// TIA Portal project "Mel7_new" (V15.1) (continued)
   L_1c_45."Уставка: Недолёт" := 4.0;
   L_1c_45.PV := 0.1030816;
   L_1c_45.Ток := 4.001736;
   L_1c_45.AnimCode := 0;
   L_1c_45.Error := 16#0000;
   L_1c_45.Bipolar := FALSE;
   L_1c_45.Overshoot_MIN := 27649;
   L_1c_45.Undershoot_MAX := -1;
END_DATA_BLOCK

DATA_BLOCK "02_DB_DI"   // DB2
{ S7_Optimized_Access := 'FALSE' }
VERSION : 0.1
BEGIN
END_DATA_BLOCK

DATA_BLOCK "03_DB_PID"   // DB3
{ S7_Optimized_Access := 'FALSE' }
VERSION : 0.1
   VAR
      PCHNasos1 : "PID_STR";
      PCHNasos2 : "PID_STR";
      PCHNasos3 : "PID_STR";
      PCHNasos4 : "PID_STR";
      PCHNasos5 : "PID_STR";
      PCHNasos6 : "PID_STR";
      PCHNasos7 : "PID_STR";
      Gaink6_1 : Real := -0.2;
      Gaink6_2 : Real := -1.0;
      Gaink6_3 : Real := -1.0;
   END_VAR
BEGIN
   PCHNasos1.SP := 22.0;
   PCHNasos1.PV := 9.6318;
   PCHNasos1.Gain := 0.2;
   PCHNasos1.Ti := T#1M_39S;
   PCHNasos1.Td := T#0MS;
   PCHNasos1.Tm_lag := T#2S;
   PCHNasos1.Man_ON := TRUE;
   PCHNasos1.MAN := 36.0;
   PCHNasos1.LMN_HI := 50.0;
   PCHNasos1.LMN_LO := 25.0;
   PCHNasos1.Reset := FALSE;
   PCHNasos1.LMN := 72.0;
   PCHNasos2.SP := 20.0;
   PCHNasos2.PV := 9.6318;
   PCHNasos2.Gain := 1.0;
   PCHNasos2.Ti := T#20S;
   PCHNasos2.Td := T#0MS;
   PCHNasos2.Tm_lag := T#2S;
   PCHNasos2.Man_ON := TRUE;
   PCHNasos2.MAN := 40.0;
   PCHNasos2.LMN_HI := 50.0;
   PCHNasos2.LMN_LO := 20.0;
   PCHNasos2.Reset := FALSE;
   PCHNasos2.LMN := 80.0;
   PCHNasos3.SP := 20.0;
   PCHNasos3.PV := 9.6318;
   PCHNasos3.Gain := 1.0;
   PCHNasos3.Ti := T#20S;
   PCHNasos3.Td := T#0MS;
   PCHNasos3.Tm_lag := T#2S;
   PCHNasos3.Man_ON := TRUE;
   PCHNasos3.MAN := 54.0;
   PCHNasos3.LMN_HI := 54.0;
   PCHNasos3.LMN_LO := 10.0;
   PCHNasos3.Reset := FALSE;
   PCHNasos3.LMN := 98.28001;
   PCHNasos4.SP := 190.0;
   PCHNasos4.PV := 1.265914;
   PCHNasos4.Gain := 0.1;
   PCHNasos4.Ti := T#21M_40S;
   PCHNasos4.Td := T#0MS;
   PCHNasos4.Tm_lag := T#2S;
   PCHNasos4.Man_ON := TRUE;
   PCHNasos4.MAN := 10.0;
   PCHNasos4.LMN_HI := 40.0;
   PCHNasos4.LMN_LO := 10.0;
   PCHNasos4.Reset := FALSE;
   PCHNasos4.LMN := 25.0;
   PCHNasos5.SP := 210.0;
   PCHNasos5.PV := 1.265914;
   PCHNasos5.Gain := 0.1;
   PCHNasos5.Ti := T#21M_40S;
   PCHNasos5.Td := T#0MS;
   PCHNasos5.Tm_lag := T#2S;
   PCHNasos5.Man_ON := FALSE;
   PCHNasos5.MAN := 28.0;
   PCHNasos5.LMN_HI := 50.0;
   PCHNasos5.LMN_LO := 10.0;
   PCHNasos5.Reset := FALSE;
   PCHNasos5.LMN := 125.0;
   PCHNasos6.SP := 40.0;
   PCHNasos6.PV := 0.0;
   PCHNasos6.Gain := 2.0;
   PCHNasos6.Ti := T#20S;
   PCHNasos6.Td := T#10S;
   PCHNasos6.Tm_lag := T#2S;
   PCHNasos6.Man_ON := TRUE;
   PCHNasos6.MAN := 0.0;
   PCHNasos6.LMN_HI := 100.0;
   PCHNasos6.LMN_LO := 0.0;
   PCHNasos6.Reset := FALSE;
   PCHNasos6.LMN := 0.0;
   PCHNasos7.SP := 0.0;
   PCHNasos7.PV := 0.0;
   PCHNasos7.Gain := 2.0;
   PCHNasos7.Ti := T#20S;
   PCHNasos7.Td := T#10S;
   PCHNasos7.Tm_lag := T#2S;
   PCHNasos7.Man_ON := TRUE;
   PCHNasos7.MAN := 0.0;
   PCHNasos7.LMN_HI := 100.0;
   PCHNasos7.LMN_LO := 0.0;
   PCHNasos7.Reset := FALSE;
   PCHNasos7.LMN := 0.0;
END_DATA_BLOCK

DATA_BLOCK "04_DB_SYSTEM"   // DB4
{ S7_Optimized_Access := 'FALSE' }
VERSION : 0.1
   VAR
      Sec_pulse : Bool;
      Trigger : Bool;
      ALW_ON : Bool := true;
   END_VAR
BEGIN
END_DATA_BLOCK

DATA_BLOCK "06_DB_MOTORS"   // DB6
{ S7_Optimized_Access := 'FALSE' }
VERSION : 0.1
   VAR
      Nas1 : "Motor_STR";
      Nas2 : "Motor_STR";
      Nas3 : "Motor_STR";
      Nas4 : "Motor_STR";
      Nas5 : "Motor_STR";
      Nas6 : "Motor_STR";
      Nas7 : "Motor_STR";
      Nas8 : "Motor_STR";
      Nas9 : "Motor_STR";
      TIMERS : Struct
         Nas1 : IEC_TIMER;
         Nas2 : IEC_TIMER;
         Nas3 : IEC_TIMER;
         Nas4 : IEC_TIMER;
         Nas5 : IEC_TIMER;
         Nas6 : IEC_TIMER;
         Nas7 : IEC_TIMER;
         Nas8 : IEC_TIMER;
         Nas9 : IEC_TIMER;
      END_STRUCT;
      SP : Struct
         Nas1 : Bool;
         Nas2 : Bool;
         Nas3 : Bool;
         Nas4 : Bool;
         Nas5 : Bool;
         Nas6 : Bool;
         Nas7 : Bool;
      END_STRUCT;
      Rab : Struct
         Nas1 : Bool;
         Nas2 : Bool;
         Nas3 : Bool;
         Nas4 : Bool;
         Nas5 : Bool;
         Nas6 : Bool;
         Nas7 : Bool;
         Nas8 : Bool;
         Nas9 : Bool;
      END_STRUCT;
   END_VAR
BEGIN
END_DATA_BLOCK

DATA_BLOCK "09_alarmdb"   // DB9
{ S7_Optimized_Access := 'FALSE' }
VERSION : 0.1
   VAR
      alarmm1 : Int;
      alarmm2 : Int;
      alarmm3 : Int;
      alarmm4 : Int;
      alarmm5 : Int;
      alarmm6 : Int;
      alarmm7 : Int;
      alarmm8 : Int;
      alarmm9 : Int;
      alarmm10 : Int;
      alarmm11 : Int;
      alarmm12 : Int;
      alarmm13 : Int;
      alarmm14 : Int;
      alarmm15 : Int;
      alarmm16 : Int;
      alarmm17 : Int;
      alarmm18 : Int;
      alarmm19 : Int;
      alarmm20 : Int;
      kvit : Bool;
      sig_kvit : Bool;
      alarm_out : Bool;
      alarm_hmi : Int;
      signal_hmi : Int;
      alarmt : Struct
         alarmt1 : Bool;
         alarmt2 : Bool;
         alarmt3 : Bool;
         alarmt4 : Bool;
         alarmt5 : Bool;
         alarmt6 : Bool;
         alarmt7 : Bool;
         alarmt8 : Bool;
         alarmt9 : Bool;
         alarmt10 : Bool;
         alarmt11 : Bool;
         alarmt12 : Bool;
         alarmt13 : Bool;
         alarmt14 : Bool;
         alarmt15 : Bool;
         alarmt16 : Bool;
         alarmt17 : Bool;
         alarmt18 : Bool;
         alarmt19 : Bool;
         alarmt20 : Bool;
      END_STRUCT;
      signal : Struct
         alarmt1 : Bool;
         alarmt2 : Bool;
         alarmt3 : Bool;
         alarmt4 : Bool;
         alarmt5 : Bool;
         alarmt6 : Bool;
         alarmt7 : Bool;
         alarmt8 : Bool;
         alarmt9 : Bool;
         alarmt10 : Bool;
         alarmt11 : Bool;
         alarmt12 : Bool;
         alarmt13 : Bool;
         alarmt14 : Bool;
         alarmt15 : Bool;
         alarmt16 : Bool;
         alarmt17 : Bool;
         alarmt18 : Bool;
         alarmt19 : Bool;
         alarmt20 : Bool;
         alarmt21 : Bool;
         alarmt22 : Bool;
         alarmt23 : Bool;
         alarmt24 : Bool;
         alarmt25 : Bool;
         alarmt26 : Bool;
         alarmt27 : Bool;
         alarmt28 : Bool;
         alarmt29 : Bool;
         alarmt30 : Bool;
         alarmt31 : Bool;
         alarmt32 : Bool;
      END_STRUCT;
   END_VAR
BEGIN
END_DATA_BLOCK

DATA_BLOCK "11_db_narabotki"   // DB11
{ S7_Optimized_Access := 'FALSE' }
VERSION : 0.1
   VAR
      Nas1_narab : "Narabotki";
      Nas2_narab : "Narabotki";
      Nas3_narab : "Narabotki";
      Nas4_narab : "Narabotki";
      Nas5_narab : "Narabotki";
   END_VAR
BEGIN
END_DATA_BLOCK

DATA_BLOCK "DB_PCHNasos1"   // DB15
{ S7_Optimized_Access := 'FALSE' }
AUTHOR : SIMATIC
FAMILY : ICONT
NAME : CONT_C
VERSION : 0.0
// stored: InstanceOfName CONT_C
"CONT_C"
BEGIN
END_DATA_BLOCK

DATA_BLOCK "DB_PCHNasos2"   // DB16
{ S7_Optimized_Access := 'FALSE' }
AUTHOR : SIMATIC
FAMILY : ICONT
NAME : CONT_C
VERSION : 0.0
// stored: InstanceOfName CONT_C
"CONT_C"
BEGIN
END_DATA_BLOCK

DATA_BLOCK "DB_PCHNasos3"   // DB17
{ S7_Optimized_Access := 'FALSE' }
AUTHOR : SIMATIC
FAMILY : ICONT
NAME : CONT_C
VERSION : 0.0
// stored: InstanceOfName CONT_C
"CONT_C"
BEGIN
END_DATA_BLOCK

DATA_BLOCK "DB_PCHNasos4"   // DB18
{ S7_Optimized_Access := 'FALSE' }
AUTHOR : SIMATIC
FAMILY : ICONT
NAME : CONT_C
VERSION : 0.0
// stored: InstanceOfName CONT_C
"CONT_C"
BEGIN
END_DATA_BLOCK

DATA_BLOCK "DB_PCHNasos5"   // DB19
{ S7_Optimized_Access := 'FALSE' }
AUTHOR : SIMATIC
FAMILY : ICONT
NAME : CONT_C
VERSION : 0.0
// stored: InstanceOfName CONT_C
"CONT_C"
BEGIN
END_DATA_BLOCK

DATA_BLOCK "DB_PCHNasos6"   // DB20
{ S7_Optimized_Access := 'FALSE' }
AUTHOR : SIMATIC
FAMILY : ICONT
NAME : CONT_C
VERSION : 0.0
// stored: InstanceOfName CONT_C
"CONT_C"
BEGIN
END_DATA_BLOCK

DATA_BLOCK "DB_PCHNasos7"   // DB21
{ S7_Optimized_Access := 'FALSE' }
AUTHOR : SIMATIC
FAMILY : ICONT
NAME : CONT_C
VERSION : 0.0
// stored: InstanceOfName CONT_C
"CONT_C"
BEGIN
END_DATA_BLOCK

FUNCTION_BLOCK "PID lean"   // FB1, LAD
{ S7_Optimized_Access := 'TRUE' }
VERSION : 0.1
   VAR_INPUT
      SP : Real := 0.0;
      PV : Real := 0.0;
      Gain : Real := 2.0;
      Ti : Time := T#20s;
      Td : Time := T#10s;
      Tm_lag : Time := T#2s;
      Man_ON : Bool := true;
      MAN : Real := 0.0;
      LMN_HI : Real := 100.0;
      LMN_LO : Real := 0.0;
      Reset : Bool;
   END_VAR
   VAR_OUTPUT
      LMN : Real := 0.0;
   END_VAR
   VAR
      IEC_Timer_0 : IEC_TIMER;
      "Last Time" : Time := T#0ms;
      IEC_Timer_1 : IEC_TIMER;
      DeltaTimeR : Real := 0.0;
      "Always On" : Bool;
      ER : Real := 0.0;
      Last_ER : Real := 0.0;
      LMN_P : Real := 0.0;
      LMN_I : Real := 0.0;
      LMN_D : Real := 0.0;
      LMN_AUTO : Real := 0.0;
   END_VAR
   VAR_TEMP
      ET : Time;
      DeltaTimeDI : DInt;
      AuxDI1 : DInt;
      AuxDI2 : DInt;
      Ti_R : Real;
      Td_R : Real;
      Tm_R : Real;
      AuxR : Real;
      AuxR2 : Real;
      DeltaER : Real;
   END_VAR
   VAR_TEMP   // added for the SCL form of the ladder/FBD networks
      _w1 : Bool;
   END_VAR
BEGIN

REGION Network 1: always on
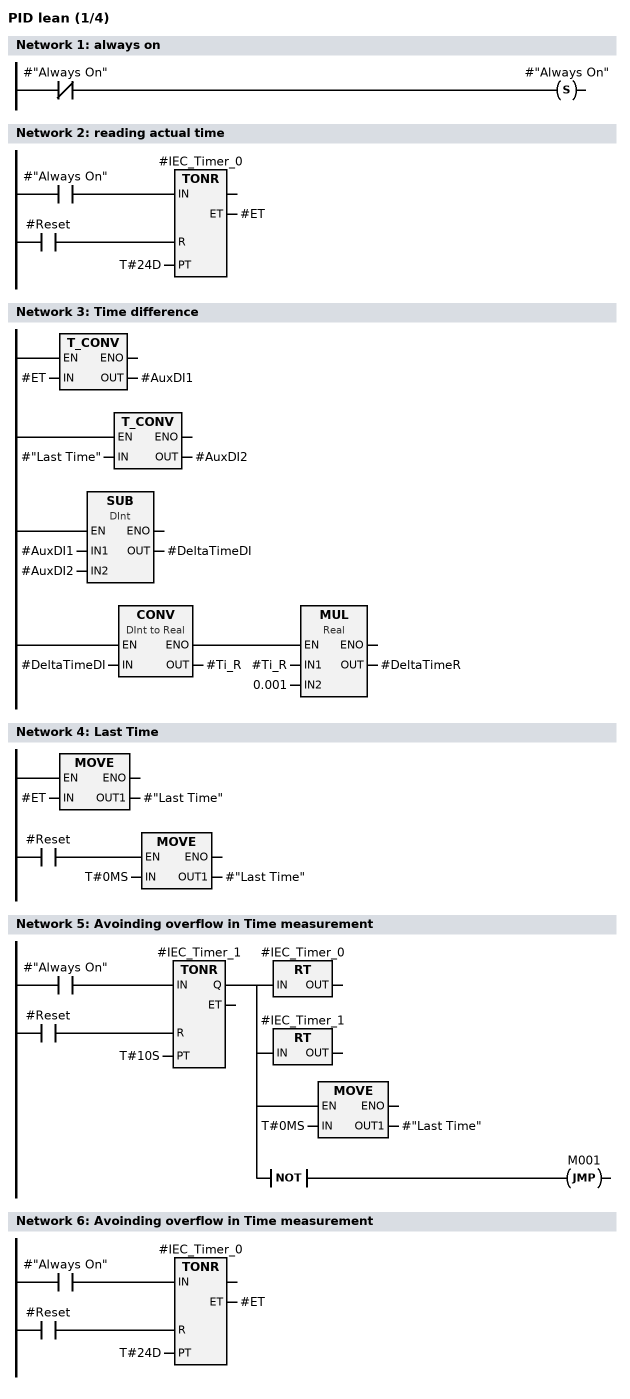
   RUNG wire#powerrail
      I_Contact( #"Always On" )
      S_Coil( #"Always On" )
   END_RUNG
   // the same network as SCL:
   IF NOT #"Always On" THEN #"Always On" := TRUE; END_IF;
END_REGION

REGION Network 2: reading actual time
   #IEC_Timer_0.TONR(IN := #"Always On", R := #Reset, PT := T#24D, ET => #ET);
END_REGION

REGION Network 3: Time difference
   // ENO of a box is taken as its EN; it also drops when the box reports an error
   #AuxDI1 := T_CONV(IN := #ET);
   #AuxDI2 := T_CONV(IN := #"Last Time");
   #DeltaTimeDI := #AuxDI1 - #AuxDI2;
   #Ti_R := DINT_TO_REAL(#DeltaTimeDI);
   #DeltaTimeR := #Ti_R * 0.001;
END_REGION

REGION Network 4: Last Time
   RUNG wire#powerrail
      { S7_GenerateENO := "TRUE" } Move(in := #ET, out1 => #"Last Time")
   END_RUNG
   RUNG wire#powerrail
      Contact( #Reset )
      { S7_GenerateENO := "TRUE" } Move(in := T#0MS, out1 => #"Last Time")
   END_RUNG
   // the same network as SCL:
   #"Last Time" := #ET;
   IF #Reset THEN #"Last Time" := T#0MS; END_IF;
END_REGION

REGION Network 5: Avoinding overflow in Time measurement
   #IEC_Timer_1.TONR(IN := #"Always On", R := #Reset, PT := T#10S);
   IF #IEC_Timer_1.Q THEN RESET_TIMER(#IEC_Timer_0); END_IF;
   #_w1 := #IEC_Timer_1.Q;
   IF #_w1 THEN
       RESET_TIMER(#IEC_Timer_1);
       #"Last Time" := T#0MS;
   END_IF;
   IF NOT #_w1 THEN GOTO M001; END_IF;
END_REGION

REGION Network 6: Avoinding overflow in Time measurement
   #IEC_Timer_0.TONR(IN := #"Always On", R := #Reset, PT := T#24D, ET => #ET);
END_REGION

REGION Network 7: Reset
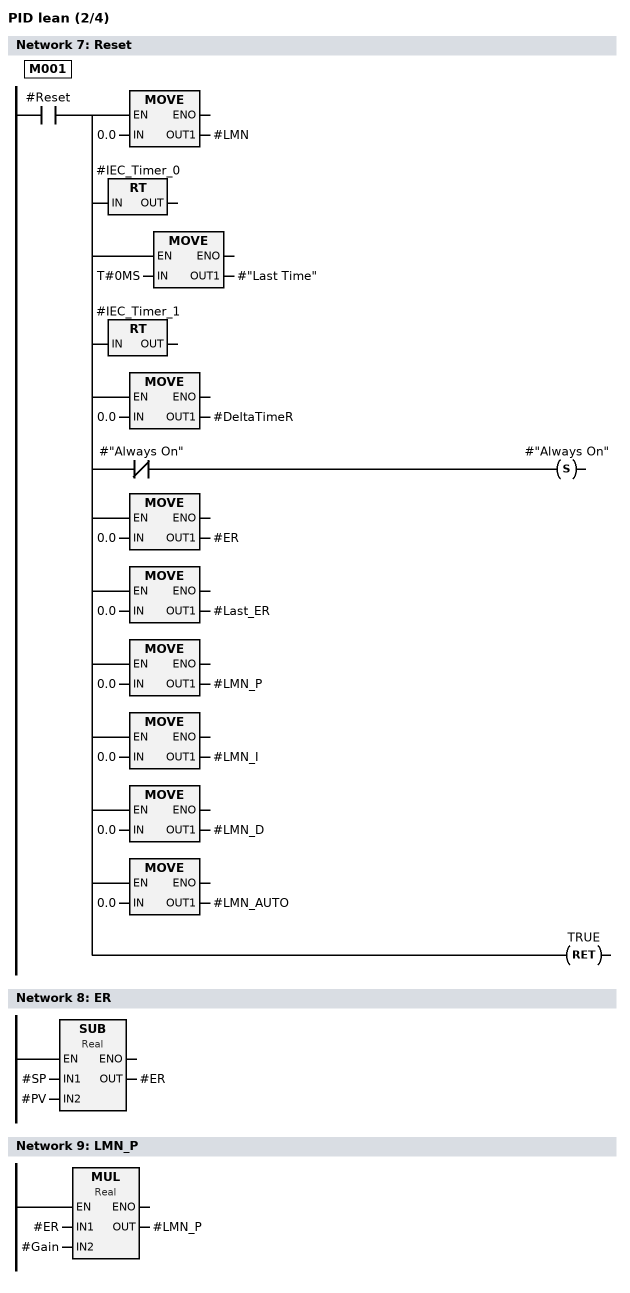
   M001:
   IF #Reset THEN
       #LMN := 0.0;
       RESET_TIMER(#IEC_Timer_0);
       #"Last Time" := T#0MS;
       RESET_TIMER(#IEC_Timer_1);
       #DeltaTimeR := 0.0;
   END_IF;
   IF #Reset AND NOT #"Always On" THEN #"Always On" := TRUE; END_IF;
   IF #Reset THEN
       #ER := 0.0;
       #Last_ER := 0.0;
       #LMN_P := 0.0;
       #LMN_I := 0.0;
       #LMN_D := 0.0;
       #LMN_AUTO := 0.0;
       ENO := TRUE;
       RETURN;
   END_IF;
END_REGION

REGION Network 8: ER
   RUNG wire#powerrail
      { S7_Templates := "SrcType := Real"; S7_GenerateENO := "TRUE" } Sub(in1 := #SP, in2 := #PV, out => #ER)
   END_RUNG
   // the same network as SCL:
   #ER := #SP - #PV;
END_REGION

REGION Network 9: LMN_P
   RUNG wire#powerrail
      { S7_Templates := "SrcType := Real"; S7_GenerateENO := "TRUE" } Mul(in1 := #ER, in2 := #Gain, out => #LMN_P)
   END_RUNG
   // the same network as SCL:
   #LMN_P := #ER * #Gain;
END_REGION

REGION Network 10: LMN_I = ER/Ti*Delta time + LMN_I
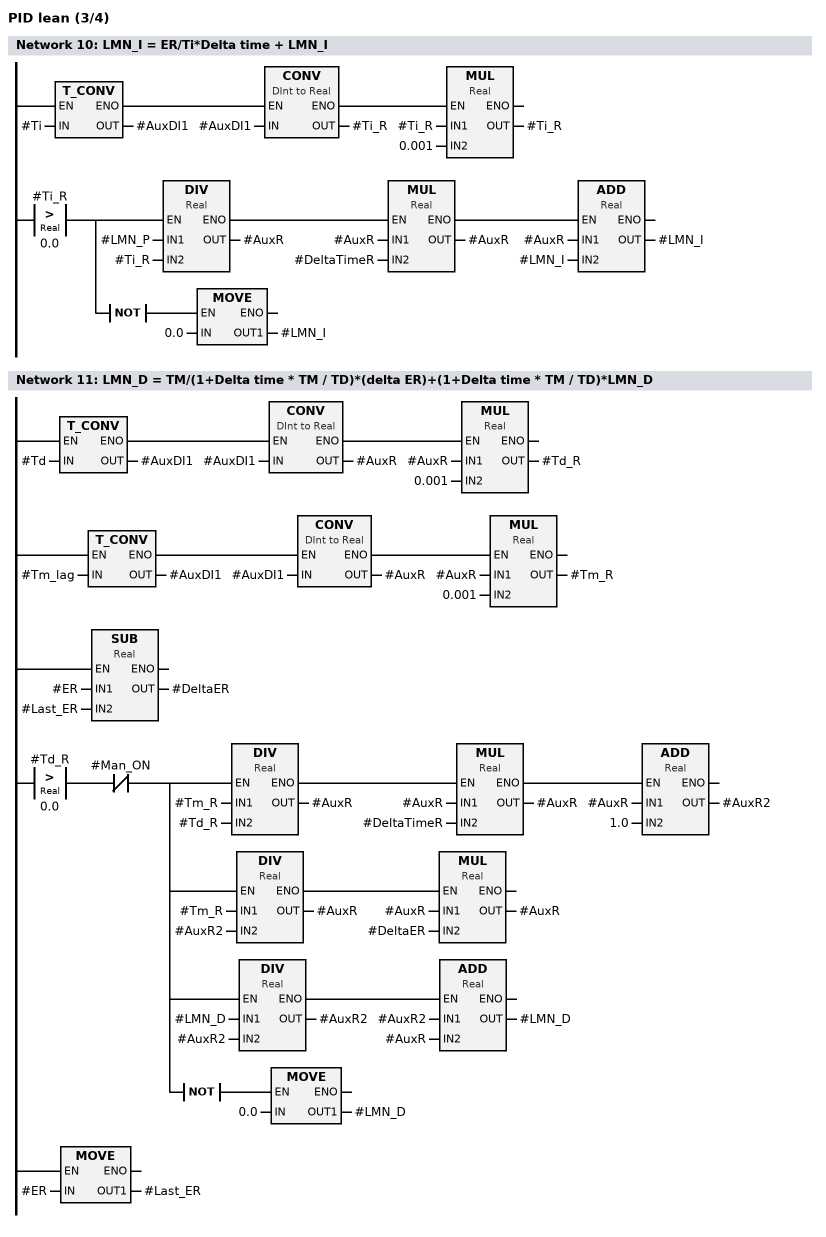
   // ENO of a box is taken as its EN; it also drops when the box reports an error
   #AuxDI1 := T_CONV(IN := #Ti);
   #Ti_R := DINT_TO_REAL(#AuxDI1);
   #Ti_R := #Ti_R * 0.001;
   #_w1 := #Ti_R > 0.0;
   IF #_w1 THEN
       #AuxR := #LMN_P / #Ti_R;
       #AuxR := #AuxR * #DeltaTimeR;
       #LMN_I := #AuxR + #LMN_I;
   END_IF;
   IF NOT #_w1 THEN #LMN_I := 0.0; END_IF;
END_REGION

REGION Network 11: LMN_D = TM/(1+Delta time * TM / TD)*(delta ER)+(1+Delta time * TM / TD)*LMN_D
   // ENO of a box is taken as its EN; it also drops when the box reports an error
   #AuxDI1 := T_CONV(IN := #Td);
   #AuxR := DINT_TO_REAL(#AuxDI1);
   #Td_R := #AuxR * 0.001;
   #AuxDI1 := T_CONV(IN := #Tm_lag);
   #AuxR := DINT_TO_REAL(#AuxDI1);
   #Tm_R := #AuxR * 0.001;
   #DeltaER := #ER - #Last_ER;
   #_w1 := (#Td_R > 0.0) AND NOT #Man_ON;
   IF #_w1 THEN
       #AuxR := #Tm_R / #Td_R;
       #AuxR := #AuxR * #DeltaTimeR;
       #AuxR2 := #AuxR + 1.0;
       #AuxR := #Tm_R / #AuxR2;
       #AuxR := #AuxR * #DeltaER;
       #AuxR2 := #LMN_D / #AuxR2;
       #LMN_D := #AuxR2 + #AuxR;
   END_IF;
   IF NOT #_w1 THEN #LMN_D := 0.0; END_IF;
   #Last_ER := #ER;
END_REGION

REGION Network 12: LMN_AUTO
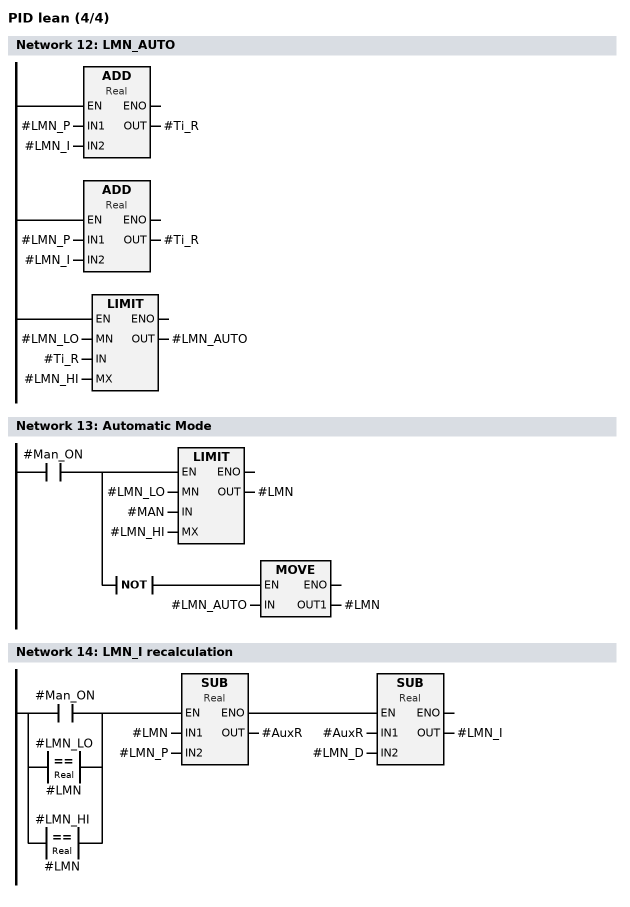
   #Ti_R := #LMN_P + #LMN_I;
   #Ti_R := #LMN_P + #LMN_I;
   #LMN_AUTO := LIMIT(MN := #LMN_LO, IN := #Ti_R, MX := #LMN_HI);
END_REGION

REGION Network 13: Automatic Mode
   IF #Man_ON THEN #LMN := LIMIT(MN := #LMN_LO, IN := #MAN, MX := #LMN_HI); END_IF;
   IF NOT #Man_ON THEN #LMN := #LMN_AUTO; END_IF;
END_REGION

REGION Network 14: LMN_I recalculation
   RUNG wire#powerrail
      Contact( #Man_ON )
      wire#w1
      { S7_Templates := "SrcType := Real"; S7_GenerateENO := "TRUE" } Sub(in1 := #LMN, in2 := #LMN_P, out => #AuxR)
      { S7_Templates := "SrcType := Real"; S7_GenerateENO := "TRUE" } Sub(in1 := #AuxR, in2 := #LMN_D, out => #LMN_I)
   END_RUNG
   RUNG wire#powerrail
      { S7_Templates := "SrcType := Real" } EQ_Contact(in1 := #LMN_LO, in2 := #LMN)
   END_RUNG wire#w1
   RUNG wire#powerrail
      { S7_Templates := "SrcType := Real" } EQ_Contact(in1 := #LMN_HI, in2 := #LMN)
   END_RUNG wire#w1
   // the same network as SCL:
   // ENO of a box is taken as its EN; it also drops when the box reports an error
   IF #Man_ON OR (#LMN_LO = #LMN) OR (#LMN_HI = #LMN) THEN
       #AuxR := #LMN - #LMN_P;
       #LMN_I := #AuxR - #LMN_D;
   END_IF;
END_REGION
END_FUNCTION_BLOCK

FUNCTION_BLOCK "CONT_C"   // FB2, SCL
{ S7_Optimized_Access := 'FALSE' }
AUTHOR : SIMATIC
FAMILY : ICONT
NAME : CONT_C
VERSION : 0.0
// reversed by komatic
   VAR_INPUT
      COM_RST : Bool;   // Полный рестарт
      MAN_ON : Bool := TRUE;   // Ручной режим включить
      PVPER_ON : Bool;   // Чтение входной переменной с периферии включить
      P_SEL : Bool := TRUE;   // Пропорциональную составляющую включить
      I_SEL : Bool := TRUE;   // Интегральную составляющую включить
      INT_HOLD : Bool;   // Удержание интегральной составляющей
      I_ITL_ON : Bool;   // Инициализировать интегральную составляющую
      D_SEL : Bool;   // Дифференциальную составляющую включить
      CYCLE : Time := T#1S;   // Время выполнения блока
      SP_INT : Real;   // Внутреннее задание
      PV_IN : Real;   // Входная переменная
      PV_PER : Word;   // Входная переменная (периферия)
      MAN : Real;   // Ручной выход
      GAIN : Real := 2.0;   // Коэффициент пропорциональности
      TI : Time := T#20S;   // Время интегрирования
      TD : Time := T#10S;   // Время дифференцирования
      TM_LAG : Time := T#2S;   // Время действия дифференциальной составляющей
      DEADB_W : Real;   // Ширина зоны нечувствительности
      LMN_HLM : Real := 100.0;   // Верхний предел выходного сигнала
      LMN_LLM : Real;   // Нижний предел выходного сигнала
      PV_FAC : Real := 1.0;   // Коэффициент для корректировки входной переменной (умножение)
      PV_OFF : Real;   // Коэффициент для корректировки входной переменной (сложение)
      LMN_FAC : Real := 1.0;   // Коэффициент для корректировки выходной переменной (умножение)
      LMN_OFF : Real;   // Коэффициент для корректировки входной переменной (сложение)
      I_ITLVAL : Real;   // Начальное значение интегральной составляющей
      DISV : Real;   // Возмущающая переменная
   END_VAR
   VAR_OUTPUT
      LMN : Real;   // Выходное значение
      LMN_PER : Word;   // Выходное значение (переферия)
      QLMN_HLM : Bool;   // Верхний предел выхода достигнут
      QLMN_LLM : Bool;   // Нижний предел выхода достигнут
      LMN_P : Real;   // Пропорциональная составляющая
      LMN_I : Real;   // Интегральная составляющая
      LMN_D : Real;   // Дифференциальная составляющая
      PV : Real;   // Входная переменная
      ER : Real;   // Сигнал рассогласования
   END_VAR
   VAR
      sInvAlt : Real;
      sIanteilAlt : Real;
      sRestInt : Real;
      sRestDif : Real;
      sRueck : Real;
      sLmn : Real;
      sbArwHLmOn : Bool;   // Выход достиг максимального значения
      sbArwLLmOn : Bool;   // Выход достиг минимального значения
      sbILimOn : Bool := TRUE;
   END_VAR
   VAR_TEMP
      Hvar : Real;   // Hilfsvariable
      rCycle : Real;   // Abtastzeit in real
      Diff : Real;   // Дnderungswert
      Istwert : Real;   // Istwert
      ErKp : Real;   // Вспомогательная переменная
      rTi : Real;   // Integrationszeit in real
      rTd : Real;   // Differentiationszeit in real
      rTmLag : Real;   // Verzцgerungszeit in real
      Panteil : Real;   // P-Anteil
      Ianteil : Real;   // I-Anteil
      Danteil : Real;   // D-Anteil
      Verstaerk : Real;   // Verstдrkung
      RueckDiff : Real;   // Differenz des Rьckkopplungswertes
      RueckAlt : Real;   // Alter Rьckkopplungswert
      dLmn : Real;   // Stellwert
      gf : Real;   // Hilfwert
      rVal : Real;   // Real Hilfsvariable
   END_VAR
BEGIN

   IF #COM_RST                                          //Полный рестарт
   THEN
       // Обнуление переменных
       #sIanteilAlt:=#I_ITLVAL;
       #LMN:=0.0;                                       //Выходное значение
       #QLMN_HLM:=0;                                    //Верхний предел выхода достигнут
       #QLMN_LLM:=0;                                    //Нижний предел выхода достигнут
       #LMN_P:=0.0;                                     //Пропорциональная составляющая
       #LMN_I:=0.0;                                     //Интегральная составляющая
       #LMN_D:=0.0;                                     //Дифференциальная составляющая
       #LMN_PER:=0;        //Выходное значение (периферия)
       #PV:=0.0;                                        //Входная переменная
       #ER:=0.0;                                        //Сигнал рассогласования
       #sInvAlt:=0.0;
       #sRestInt:=0.0;
       #sRestDif:=0.0;
       #sRueck:=0.0;
       #sLmn:=0.0;
       #sbArwHLmOn:=0;
       #sbArwLLmOn:=0;
   ELSE
       #rCycle:= DINT_TO_REAL(TIME_TO_DINT(#CYCLE)) / 1000.0;            //Время выполнения блока в секундах
       #Istwert:=INT_TO_REAL(WORD_TO_INT(#PV_PER)) * 100.0 / 27648.0;    // Получили входную переменную от периферии (0-2768 в 0-100)
       #Istwert:=#Istwert * #PV_FAC + #PV_OFF;                             // Скорректировали входную переменную
       IF NOT #PVPER_ON THEN #Istwert:=#PV_IN; END_IF;                    // Если периферийный вход отключен берем переменную из PV_IN
       #PV:= #Istwert;                                                   // Входная переменная
       #ErKp:=#SP_INT - #PV;                                              // Получили рассогласование между заданием и входом
       IF     #ErKp < (-#DEADB_W)     THEN #ER:=#ErKp+#DEADB_W;             // Если рассогласование больше зоны нечувствительности
       ELSIF  #ErKp >   #DEADB_W      THEN #ER:=#ErKp-#DEADB_W;             // уменьшаем рассогласование на величину зоны нечуств.
       ELSE                              #ER:=0.0;                      // иначе принимаем рассогласование равным нулю.
       END_IF;
       #ErKp:=#ER * #GAIN;                                                // Рассогласование, умноженное на кфт пропорциональности
       #rTi:=DINT_TO_REAL(TIME_TO_DINT(#TI)) / 1000.0;                   // Время интегрирования в секундах
       #rTd:=DINT_TO_REAL(TIME_TO_DINT(#TD)) / 1000.0;                   // Время дифференцирования в секундах
       #rTmLag:=DINT_TO_REAL(TIME_TO_DINT(#TM_LAG)) / 1000.0;            // Время действия диф.составляющей в секундах
       // Проверка на допустимость временных настроек регулятора
       IF #rTi < (#rCycle * 0.5)     THEN    #rTi:=#rCycle * 0.5;      END_IF; // Минимальное время интегрирования - Cycle / 2
       IF #rTd < #rCycle             THEN    #rTd:=#rCycle;            END_IF; // Минимальное время дифференцирования - Cycle
       IF #rTmLag < #rCycle * 0.5    THEN    #rTmLag:=#rCycle * 0.5;   END_IF; // Минимальное время действия диф.сост.- Cycle / 2
       // Вычисление пропорциональной составляющей
       IF #P_SEL
       THEN
           #Panteil:=#ErKp;                                              // Если выбрана пропорциональная составляющая
       ELSE
           #Panteil:=0.0;
       END_IF;
       //---------------------------------------------------------------------------------------------
       // Вычисление интегральной составляющей
       //---------------------------------------------------------------------------------------------   
       IF #I_SEL                    //Интегральную составляющую включить
       THEN
           IF #I_ITL_ON             //Инициализировать интегральную составляющую
           THEN
               #Ianteil:=#I_ITLVAL;
               #sRestInt:=0.0;
           ELSE
               IF #MAN_ON           //Ручной режим
               THEN
                   #Ianteil:=#sLmn - #Panteil - #DISV;
                   #sRestInt:=0.0;
               ELSE                //Автоматический режим
                   #Diff:=#rCycle / #rTi *(#ErKp + #sInvAlt) *  0.5 + #sRestInt;
                   IF ((#Diff>0.0) AND #sbArwHLmOn OR #INT_HOLD)OR ((#Diff<0.0) AND #sbArwLLmOn) THEN #Diff:=0.0; END_IF;       
                   #Ianteil:=#sIanteilAlt + #Diff;
                   #sRestInt:=#sIanteilAlt - #Ianteil + #Diff;
               END_IF;
           END_IF;
       ELSE
           #Ianteil:=0.0;
           #sRestInt:=0.0;
       END_IF;
       //---------------------------------------------------------------------------------------------
       //Формирование дифференциальной составляющей
       //---------------------------------------------------------------------------------------------   
       #Diff:=#ErKp;
       IF (NOT #MAN_ON) AND #D_SEL
       THEN
           #Verstaerk:= #rTd / (#rCycle * 0.5 + #rTmLag);
           #Danteil:= (#Diff - #sRueck) * #Verstaerk;
           #RueckAlt:= #sRueck;
           #RueckDiff:= #rCycle / #rTd * #Danteil + #sRestDif;
           #sRueck:= #RueckDiff + #RueckAlt;
           #sRestDif:=#RueckAlt - #sRueck + #RueckDiff;
       ELSE
           #Danteil:=0.0;   
           #sRestDif:=0.0;
           #sRueck:=#Diff;
       END_IF;
       //---------------------------------------------------------------------------------------------
       //Формирование выхода
       //---------------------------------------------------------------------------------------------
       #dLmn:=#Panteil + #Ianteil + #Danteil + #DISV;
       IF #MAN_ON           // Если ручной режим
       THEN
           #dLmn:=#MAN;      // Ручной выход
       ELSE
           IF (NOT #I_ITL_ON) AND #I_SEL
           THEN
               IF (#Ianteil > (#LMN_HLM - #DISV)) AND (#dLmn > #LMN_HLM) AND ((#dLmn - #LMN_D)> #LMN_HLM)
               THEN
                   #rVal:=#LMN_HLM - #DISV;
                   #gf:=  #dLmn - #LMN_HLM;
                   #rVal:=#Ianteil - #rVal;
                   IF  #rVal > #gf THEN #rVal:=#gf; END_IF;
                   #Ianteil:=#Ianteil - #rVal;
               ELSE
                   IF (#Ianteil < (#LMN_LLM - #DISV)) AND (#dLmn < #LMN_LLM) AND ((#dLmn - #LMN_D) < #LMN_LLM)
                   THEN
                       #rVal:=#LMN_LLM - #DISV;
                       #gf:=#dLmn - #LMN_LLM;
                       #rVal:=#Ianteil - #rVal;
                       IF #rVal < #gf  THEN #rVal:=#gf; END_IF;
                       #Ianteil:=#Ianteil - #rVal;
                   END_IF;   
                END_IF;      
           END_IF;
       END_IF;
       #LMN_P:=#Panteil;
       #LMN_I:=#Ianteil;
       #LMN_D:=#Danteil;
       #sInvAlt:=#ErKp;
       #sIanteilAlt:=#Ianteil;
       #sbArwHLmOn:=0;
       #sbArwLLmOn:=0;
       IF (#dLmn >= #LMN_HLM)
       THEN
           #QLMN_HLM:=1;
           #QLMN_LLM:=0;
           #dLmn:=#LMN_HLM;
           #sbArwHLmOn:=1;
       ELSE
           #QLMN_HLM:=0;
           IF (#dLmn <= #LMN_LLM)
           THEN
               #QLMN_LLM:=1;
               #dLmn:=#LMN_LLM;
               #sbArwLLmOn:=1;
           ELSE
               #QLMN_LLM:=0; 
           END_IF;
       END_IF;
       #sLmn:=#dLmn;
       #dLmn:=#sLmn * #LMN_FAC + #LMN_OFF;  
       #LMN:=#dLmn;
       #dLmn:=#LMN * 2.764800e+002;
       IF #dLmn >= 3.251100e+004
       THEN
           #dLmn:=3.251100e+004;
       ELSE
           IF #dLmn <= -3.251200e+004
           THEN
               #dLmn:=-3.251200e+004;
           END_IF;
       END_IF;
       #LMN_PER:= INT_TO_WORD(REAL_TO_INT(#dLmn));
   END_IF;
END_FUNCTION_BLOCK

FUNCTION_BLOCK "CONT_S"   // FB3, SCL
{ S7_Optimized_Access := 'FALSE' }
VERSION : 0.0
// reversed by komatic
   VAR_INPUT
      COM_RST : Bool;   // полный рестарт
      LMNR_HS : Bool;   // high limit signal of repeated manipulated value
      LMNR_LS : Bool;   // low limit signal of repeated manipulated value
      LMNS_ON : Bool;   // manipulated signals on
      LMNUP : Bool;   // manipulated signal up
      LMNDN : Bool;   // manipulated signal down
      PVPER_ON : Bool;   // брать входную переменную из периферии
      CYCLE : Time := T#1S;   // время выполнения блока
      SP_INT : Real;   // внутреннее задание
      PV_IN : Real;   // входная переменная
      PV_PER : Word;   // входная переменная, периферия
      GAIN : Real := 2.0;   // кфт пропорциональности
      TI : Time := T#20S;   // время интегрирования
      DEADB_W : Real := 1.0;   // dead band width
      PV_FAC : Real := 1.0;   // масштабирующий кфт входной переменной
      PV_OFF : Real;   // суммирующий кфт входной переменной
      PULSE_TM : Time := T#3S;   // minimum pulse time
      BREAK_TM : Time := T#3S;   // minimum break time
      MTR_TM : Time := T#30S;   // motor manipulated value
      DISV : Real;   // возмущающее воздействие
   END_VAR
   VAR_OUTPUT
      QLMNUP : Bool;   // manipulated signal up
      QLMNDN : Bool;   // manipulated signal down
      PV : Real;   // process variable
      ER : Real;   // error signal
   END_VAR
   VAR
      LMNRS_ON : Bool;
      LMNRSVAL : Real;
      LMNR_SIM : Real;
      sFbPVal : Real;
      sThrOn : Real;
      siImpAus : Int;
      stImpDauer : Time;
      stPausDauer : Time;
   END_VAR
   VAR_TEMP
      Hvar : Real;   // вспомогательная переменная
      rCycle : Real;   // Abtastzeit in real
      Istwert : Real;   // Istwert
      ErKp : Real;   // вспомогательная переменная
      rTi : Real;   // время интегрирования в real
      AdapIn1 : Real;   // Eingang 1 der Adaption der Ansprechschwelle
      AdapIn2 : Real;   // Eingang 2 der Adaption der Ansprechschwelle
      iImpEin : Int;   // Eingang des Impulsformers
      rMtrTm : Real;   // Motorstellzeit in real
      rThrOff : Real;   // Abschaltschwelle
      dInteg : Real;   // Eingang des Integrierers in der Rьckfьhrung
      dThrStIn : Real;   // three-step element input
      LmnrSim : Real;   // simulierte Stellungsrьckmeldung
   END_VAR
BEGIN

